(* Logix 5000 project; controller PLC_MCC1201_220AP1 vendor 1 type 14 code 164 rev 35.11; software revision 35.00; part 2 of 25 *)
(* tags used below, declared in another part *)
   N124 : DINT[414];
   N125 : DINT[414];
   N15 : DINT[1000];
   N179 : DINT[600];
   N251 : DINT[999];
   N42 : DINT[89];
   N43 : DINT[240];
   N45 : DINT[58];
   N46 : DINT[7];
   N54 : DINT[501];
   N60 : DINT[420];
   N61 : DINT[100];
   N7 : DINT[250];
   N98 : DINT[20];
   O : INT[128];
   S : INT[128];
   Status : INT;   // INT tag to retrieve Status value through GSV created during conversion
   T4 : TIMER[100];
   T51 : TIMER[13];
   TONY : ALIAS FOR B3[10].15;
   W_N7 : DINT[933];

ADD_ON_INSTRUCTION AOI_AccessArea_Logic   (* revision 1.0, vendor Bottero *)
// Help:
// (AOI_AccessArea_Logic,IN_xResetAlarm,IN_xEnableControlError,IN_xCycleON,IN_xConditionOkAccessArea,IN_xPhaseInProgressArea,IN_xExternalConditionOkToWork,IN_xSBRequestAccessAreaSelector,IN_xSBRequestAccessAreaButton,IN_xSBResetAccessArea,IN_xSBInternalResetArea,IN_xStatusDoorPH,IN_xSafetyOk,IN_xLampClock,tHMR,tAlm);
VAR_IN_OUT
   tAlm : AOI_AccessArea_Alm; {required}
   tHMR : AOI_AccessArea_HMR; {required}
END_VAR
VAR_INPUT
   IN_xConditionOkAccessArea : BOOL; {access None}
   IN_xCycleON : BOOL; {access None}
   IN_xEnableControlError : BOOL; {access None}
   IN_xLampClock : BOOL; {access None}
   IN_xPhaseInProgressArea : BOOL; {access None}
   IN_xResetAlarm : BOOL; {access None}
   IN_xSafetyOk : BOOL; {access None}
   IN_xSBInternalResetArea : BOOL; {access None}
   IN_xSBRequestAccessAreaButton : BOOL; {access None}
   IN_xSBRequestAccessAreaSelector : BOOL; {access None}
   IN_xSBResetAccessArea : BOOL; {access None}
   IN_xStatusDoorPH : BOOL; {access None}
END_VAR
VAR_OUTPUT
   OUT_xAccessAreaAccepted : BOOL; {access None}
   OUT_xAccessAreaRequest : BOOL; {access None}
   OUT_xConditionOkToWork : BOOL; {access None}
   OUT_xReqResetPhase : BOOL; {access None}
   OUT_xReqResetSafetyArea : BOOL; {access None}
   OUT_xSafetyAreaIntervened : BOOL;
   OUT_xSBLampAccessArea : BOOL;
   OUT_xSBLampInternalReset : BOOL;
   OUT_xSQOpeningDoor : BOOL;
   OUT_xStopFault : BOOL; {access None}
END_VAR
VAR_INPUT
   IN_xSAEnableResetAreaSafety : BOOL; {access None}
END_VAR
VAR
   tAOI_AccessArea_GP : AOI_AccessArea; {access None}
   ST_xConditionOkForceAccess : BOOL; {access None}
   ST_xConditionOkForRequestAccessArea : BOOL; {access None}
   ST_xErrorMutingDuringAccessArea : BOOL; {access None}
   ST_xFault : BOOL; {access None}
   ST_xInternalResetAreaRequired : BOOL; {access None}
   ST_xRequestResetPhase : BOOL; {access None}
   ST_xRequestResetSafetyArea : BOOL; {access None}
   ST_xStopFault : BOOL; {access None}
   ST_xWarning : BOOL; {access None}
   tm_ErrorMutingDuringAccessArea : TIMER; {access None}
   TMP_dAlarm : DINT; {access None}
   InitAlm : UDT_Spare32bit_Alm; {access None}
END_VAR

ROUTINE Logic   (* ladder *)
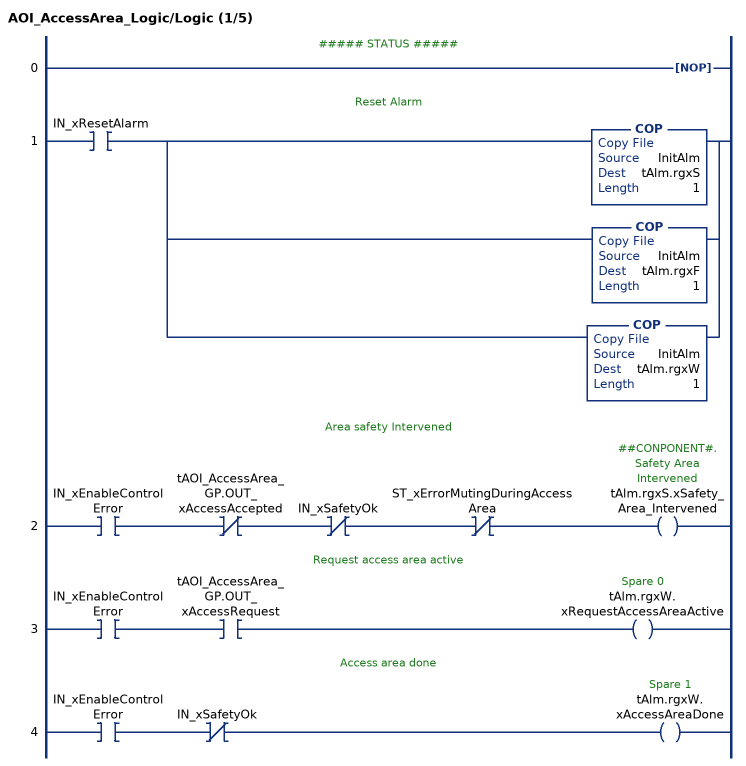
   // ##### STATUS #####
   0: NOP();
   // Reset Alarm
   1: XIC(IN_xResetAlarm)[COP(InitAlm,tAlm.rgxS,1) ,COP(InitAlm,tAlm.rgxF,1) ,COP(InitAlm,tAlm.rgxW,1) ];
   // Area safety Intervened
   2: XIC(IN_xEnableControlError)XIO(tAOI_AccessArea_GP.OUT_xAccessAccepted)XIO(IN_xSafetyOk)XIO(ST_xErrorMutingDuringAccessArea)OTE(tAlm.rgxS.xSafety_Area_Intervened);
   // Request access area active
   3: XIC(IN_xEnableControlError)XIC(tAOI_AccessArea_GP.OUT_xAccessRequest)OTE(tAlm.rgxW.xRequestAccessAreaActive);
   // Access area done
   4: XIC(IN_xEnableControlError)XIO(IN_xSafetyOk)OTE(tAlm.rgxW.xAccessAreaDone);
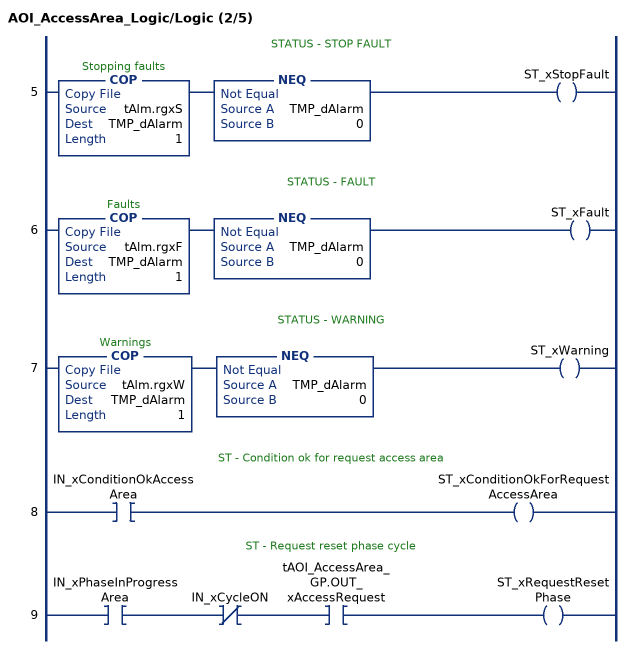
   // STATUS - STOP FAULT
   5: COP(tAlm.rgxS,TMP_dAlarm,1)NEQ(TMP_dAlarm,0)OTE(ST_xStopFault);
   // STATUS - FAULT
   6: COP(tAlm.rgxF,TMP_dAlarm,1)NEQ(TMP_dAlarm,0)OTE(ST_xFault);
   // STATUS - WARNING
   7: COP(tAlm.rgxW,TMP_dAlarm,1)NEQ(TMP_dAlarm,0)OTE(ST_xWarning);
   // ST - Condition ok for request access area
   8: XIC(IN_xConditionOkAccessArea)OTE(ST_xConditionOkForRequestAccessArea);
   // ST - Request reset phase cycle
   9: XIC(IN_xPhaseInProgressArea)XIO(IN_xCycleON)XIC(tAOI_AccessArea_GP.OUT_xAccessRequest)OTE(ST_xRequestResetPhase);
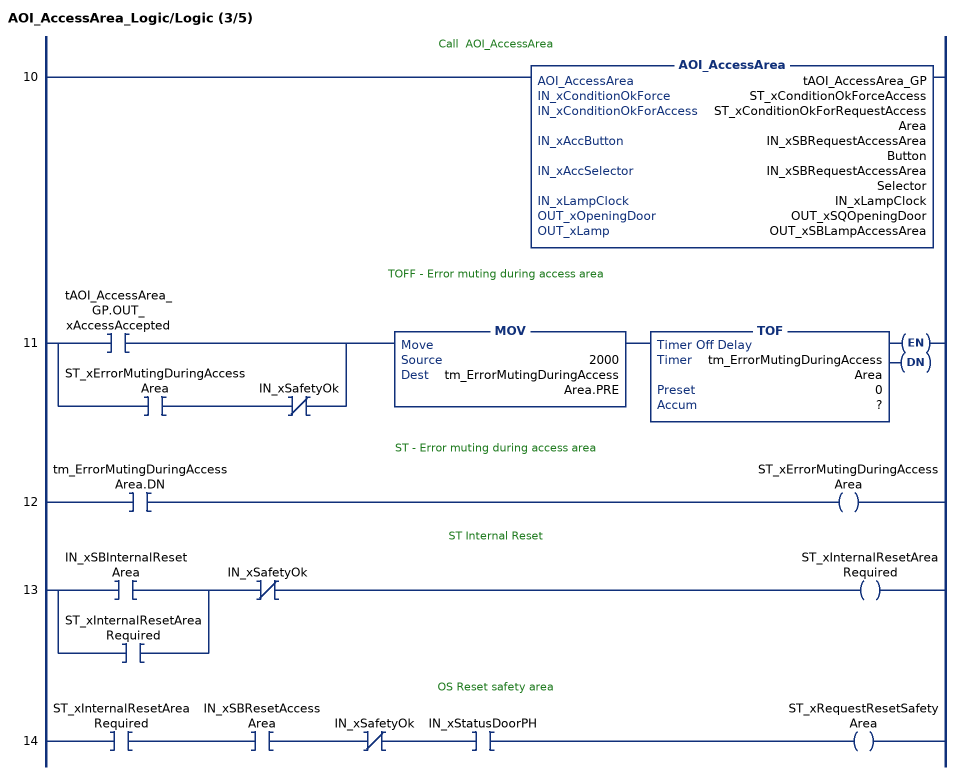
   // Call  AOI_AccessArea
   10: AOI_AccessArea(tAOI_AccessArea_GP,ST_xConditionOkForceAccess,ST_xConditionOkForRequestAccessArea,IN_xSBRequestAccessAreaButton,IN_xSBRequestAccessAreaSelector,IN_xLampClock,OUT_xSQOpeningDoor,OUT_xSBLampAccessArea);
   // TOFF - Error muting during access area
   11: [XIC(tAOI_AccessArea_GP.OUT_xAccessAccepted) ,XIC(ST_xErrorMutingDuringAccessArea) XIO(IN_xSafetyOk) ]MOV(2000,tm_ErrorMutingDuringAccessArea.PRE)TOF(tm_ErrorMutingDuringAccessArea,?,?);
   // ST - Error muting during access area
   12: XIC(tm_ErrorMutingDuringAccessArea.DN)OTE(ST_xErrorMutingDuringAccessArea);
   // ST Internal Reset
   13: [XIC(IN_xSBInternalResetArea) ,XIC(ST_xInternalResetAreaRequired) ]XIO(IN_xSafetyOk)OTE(ST_xInternalResetAreaRequired);
   // OS Reset safety area
   14: XIC(ST_xInternalResetAreaRequired)XIC(IN_xSBResetAccessArea)XIO(IN_xSafetyOk)XIC(IN_xStatusDoorPH)OTE(ST_xRequestResetSafetyArea);
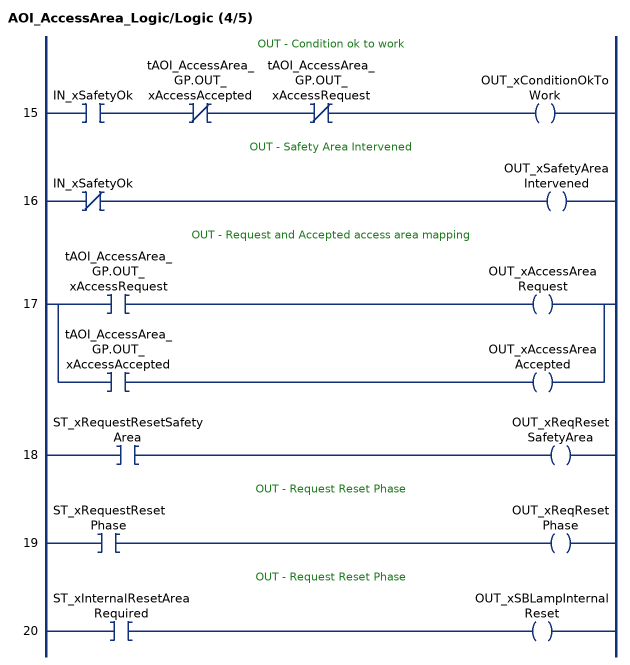
   // OUT - Condition ok to work
   15: XIC(IN_xSafetyOk)XIO(tAOI_AccessArea_GP.OUT_xAccessAccepted)XIO(tAOI_AccessArea_GP.OUT_xAccessRequest)OTE(OUT_xConditionOkToWork);
   // OUT - Safety Area Intervened
   16: XIO(IN_xSafetyOk)OTE(OUT_xSafetyAreaIntervened);
   // OUT - Request and Accepted access area mapping
   17: [XIC(tAOI_AccessArea_GP.OUT_xAccessRequest) OTE(OUT_xAccessAreaRequest) ,XIC(tAOI_AccessArea_GP.OUT_xAccessAccepted) OTE(OUT_xAccessAreaAccepted) ];
   18: XIC(ST_xRequestResetSafetyArea)OTE(OUT_xReqResetSafetyArea);
   // OUT - Request Reset Phase
   19: XIC(ST_xRequestResetPhase)OTE(OUT_xReqResetPhase);
   // OUT - Request Reset Phase
   20: XIC(ST_xInternalResetAreaRequired)OTE(OUT_xSBLampInternalReset);
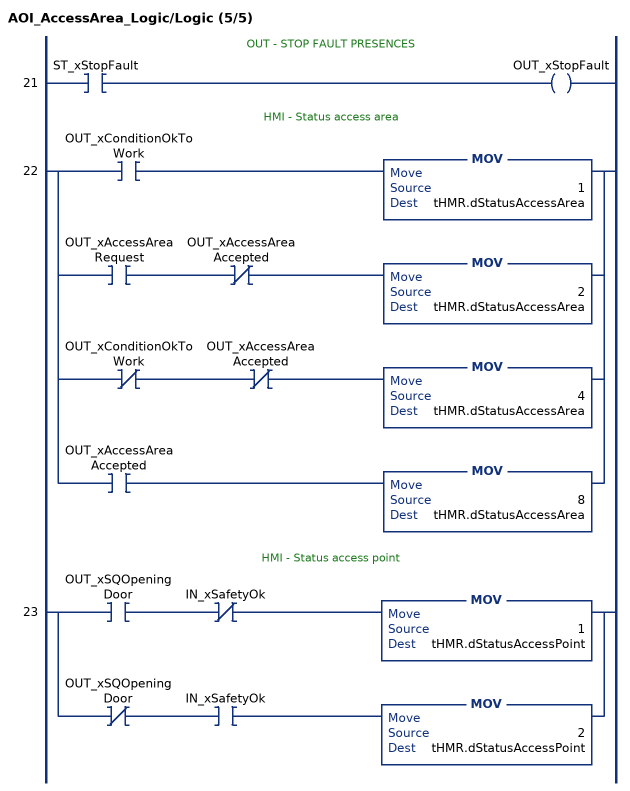
   // OUT - STOP FAULT PRESENCES
   21: XIC(ST_xStopFault)OTE(OUT_xStopFault);
   // HMI - Status access area
   22: [XIC(OUT_xConditionOkToWork) MOV(1,tHMR.dStatusAccessArea) ,XIC(OUT_xAccessAreaRequest) XIO(OUT_xAccessAreaAccepted) MOV(2,tHMR.dStatusAccessArea) ,XIO(OUT_xConditionOkToWork) XIO(OUT_xAccessAreaAccepted) MOV(4,tHMR.dStatusAccessArea) ,XIC(OUT_xAccessAreaAccepted) MOV(8,tHMR.dStatusAccessArea) ];
   // HMI - Status access point
   23: [XIC(OUT_xSQOpeningDoor) XIO(IN_xSafetyOk) MOV(1,tHMR.dStatusAccessPoint) ,XIO(OUT_xSQOpeningDoor) XIC(IN_xSafetyOk) MOV(2,tHMR.dStatusAccessPoint) ];
END_ROUTINE
END_ADD_ON_INSTRUCTION

ADD_ON_INSTRUCTION GP_AccessArea   (* revision 1.0 *)
VAR_IN_OUT
   STC : GP_AccessArea_STC; {required}
END_VAR
VAR_INPUT
   IN_xAccSelector : BOOL; {access None, required}
   IN_xAccButton : BOOL; {access None, required}
   IN_xConditionOkAccess : BOOL; {access None, required}
   IN_xConditionOkForcedAccess : BOOL; {access None, required}
   IN_xLampClock : BOOL; {access None, required}
END_VAR
VAR_OUTPUT
   OUT_xOpeningDoor : BOOL; {access None}
   OUT_xLamp : BOOL; {access None, required}
END_VAR

ROUTINE Logic   (* ladder *)
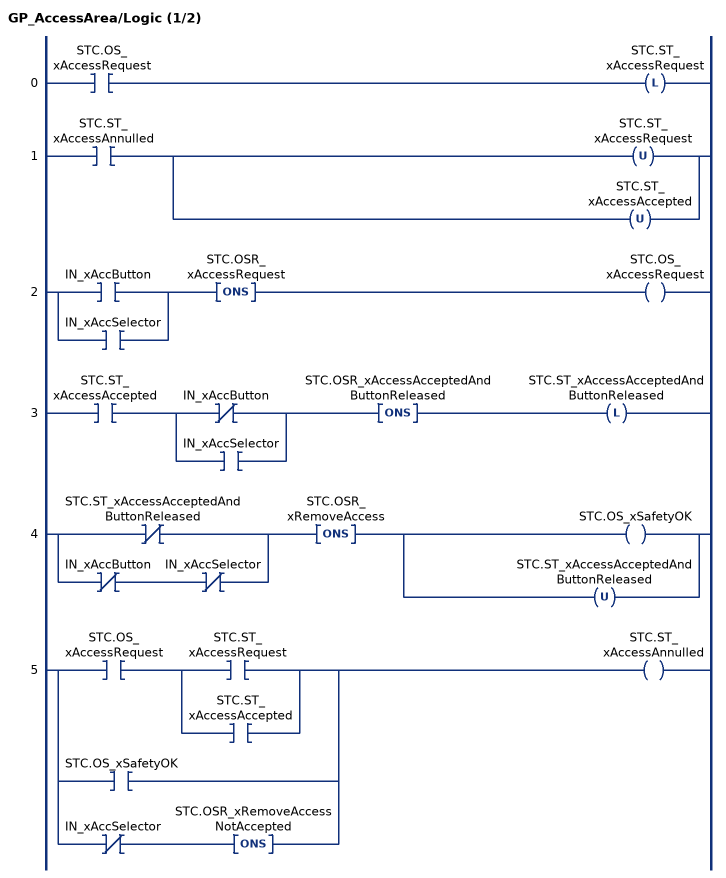
   0: XIC(STC.OS_xAccessRequest)OTL(STC.ST_xAccessRequest);
   1: XIC(STC.ST_xAccessAnnulled)[OTU(STC.ST_xAccessRequest) ,OTU(STC.ST_xAccessAccepted) ];
   2: [XIC(IN_xAccButton) ,XIC(IN_xAccSelector) ]ONS(STC.OSR_xAccessRequest)OTE(STC.OS_xAccessRequest);
   3: XIC(STC.ST_xAccessAccepted)[XIO(IN_xAccButton) ,XIC(IN_xAccSelector) ]ONS(STC.OSR_xAccessAcceptedAndButtonReleased)OTL(STC.ST_xAccessAcceptedAndButtonReleased);
   4: [XIO(STC.ST_xAccessAcceptedAndButtonReleased) ,XIO(IN_xAccButton) XIO(IN_xAccSelector) ]ONS(STC.OSR_xRemoveAccess)[OTE(STC.OS_xSafetyOK) ,OTU(STC.ST_xAccessAcceptedAndButtonReleased) ];
   5: [XIC(STC.OS_xAccessRequest) [XIC(STC.ST_xAccessRequest) ,XIC(STC.ST_xAccessAccepted) ] ,XIC(STC.OS_xSafetyOK) ,XIO(IN_xAccSelector) ONS(STC.OSR_xRemoveAccessNotAccepted) ]OTE(STC.ST_xAccessAnnulled);
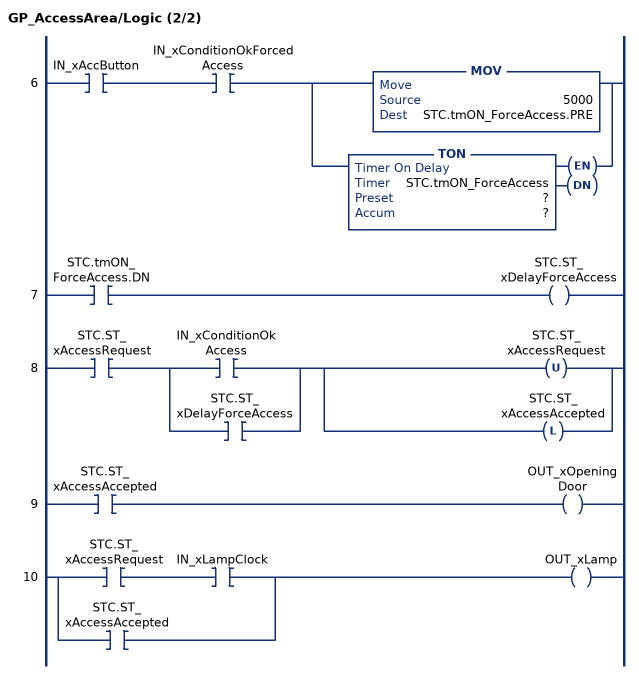
   6: XIC(IN_xAccButton)XIC(IN_xConditionOkForcedAccess)[MOV(5000,STC.tmON_ForceAccess.PRE) ,TON(STC.tmON_ForceAccess,?,?) ];
   7: XIC(STC.tmON_ForceAccess.DN)OTE(STC.ST_xDelayForceAccess);
   8: XIC(STC.ST_xAccessRequest)[XIC(IN_xConditionOkAccess) ,XIC(STC.ST_xDelayForceAccess) ][OTU(STC.ST_xAccessRequest) ,OTL(STC.ST_xAccessAccepted) ];
   9: XIC(STC.ST_xAccessAccepted)OTE(OUT_xOpeningDoor);
   10: [XIC(STC.ST_xAccessRequest) XIC(IN_xLampClock) ,XIC(STC.ST_xAccessAccepted) ]OTE(OUT_xLamp);
END_ROUTINE
END_ADD_ON_INSTRUCTION

ADD_ON_INSTRUCTION GP_NetworkDiag   (* revision 1.0 *)
VAR_IN_OUT
   IN_OB_Initialize : GP_OB_Initialize; {required}
   IN_ModuleName : MODULE; {required}   // Module name
   OUT_tModuleInfo : GP_NetworkDiag_v1; {required}   // Module info
END_VAR
VAR
   TMP_xFaulted : BOOL; {access None}
   TMP_xConnected : BOOL; {access None}
END_VAR

ROUTINE Logic   (* structured text *)
   //Initialize
   TMP_xConnected:=0;
   TMP_xFaulted:=0;
   
   //Get system info from module
   gsv(Module,IN_ModuleName,EntryStatus,OUT_tModuleInfo.dEntryStatus);
   gsv(Module,IN_ModuleName,FaultCode,OUT_tModuleInfo.dFaultCode);
   gsv(Module,IN_ModuleName,FaultInfo,OUT_tModuleInfo.dFaultInfo);
   gsv(Module,IN_ModuleName,Instance,OUT_tModuleInfo.dInstance);
   
   CASE OUT_tModuleInfo.dEntryStatus OF
   	16#0000:(*Standby: the controller is powering up.*)
    			TMP_xFaulted:= IN_OB_Initialize.OUT_xClock_800ms;
   
   	16#1000:(*Faulted: any of the MODULE object’s connections to the associated module fail.
   			This value should not be used to determine if the module failed because the MODULE
   			object leaves this state periodically when trying to reconnect to the module.
   			Instead, test for Running state (16#4000). Check for FaultCode not equal to 0 to determine if a module is faulted.
   			When Faulted, the FaultCode and FaultInfo attributes are valid until the fault condition is corrected.*)
    			TMP_xConnected:= IN_OB_Initialize.OUT_xClock_1s;
   			TMP_xFaulted:= 1;
   
   	16#2000:(*Validating: the MODULE object is verifying MODULE object integrity prior to establishing connections to the module.*)
    			TMP_xConnected:= IN_OB_Initialize.OUT_xClock_400ms;
   
   	16#3000:(*Connecting: the MODULE object is initiating connections to the module.*)
   			TMP_xConnected:= IN_OB_Initialize.OUT_xClock_400ms;
   
   	16#4000:(*Running: all connections to the module are established and data is successfully transferring.*)
    			TMP_xConnected:= 1;
   
   	16#5000:(*Shutting down: the MODULE object is in the process of shutting down all connections to the module.*)
   			TMP_xConnected:= IN_OB_Initialize.OUT_xClock_1s;
   
   	16#6000:(*Inhibited: the MODULE object is inhibited (the inhibit bit in the Mode attribute is set).*)
    			TMP_xConnected:= IN_OB_Initialize.OUT_xClock_1s;
   
   	16#7000:(*Waiting: the parent MODULE object upon which this MODULE object depends is not running*)
   			TMP_xConnected:= IN_OB_Initialize.OUT_xClock_1s;
   
   	16#9000:(*FirmwareUpdating: Firmware supervisor is attempting to flash the module. *)
    			TMP_xConnected:= IN_OB_Initialize.OUT_xClock_800ms;
   
   	16#A000:(*Configuring: Controller is downloading configuration to the module.
   			Either ?forward open? or (ADC) download occur during this state.*)
   			TMP_xConnected:= IN_OB_Initialize.OUT_xClock_800ms;
   END_CASE;
   
   IF OUT_tModuleInfo.dFaultCode<>0 THEN
   	TMP_xFaulted:= 1;
   	TMP_xConnected:= 0;
   END_IF;
   
   //Save status bit
   OUT_tModuleInfo.xConnected:=TMP_xConnected;
   OUT_tModuleInfo.xFaulted:=TMP_xFaulted;
   
   
   
   
   
   
   
   
   
   
   
   
   
   
   
   
   
   
   
   
END_ROUTINE
END_ADD_ON_INSTRUCTION

ADD_ON_INSTRUCTION GP_OB_Initialize   (* revision 1.0 *)
VAR_IN_OUT
   STC : GP_OB_Initialize_STC; {required}
END_VAR
VAR_INPUT
   IN_xInitialize : BOOL; {access None, required}   // Initialize values (Restart call)
END_VAR
VAR_OUTPUT
   OUT_dExecutionTime_ms : DINT; {access None}   // OB Execution time [ms]
   OUT_dMinExecutionTime_ms : DINT; {access None}   // OB Minimum execution time [ms]
   OUT_dMaxExecutionTime_ms : DINT; {access None}   // OB Maximum execution time [ms]
   OUT_xOs_100ms : BOOL; {access None}   // OS each 100ms
   OUT_xOs_200ms : BOOL; {access None}   // OS each 200ms
   OUT_xOs_400ms : BOOL; {access None}   // OS each 400ms
   OUT_xOs_500ms : BOOL; {access None}   // OS each 500ms
   OUT_xOs_800ms : BOOL; {access None}   // OS each 800ms
   OUT_xOs_1s : BOOL; {access None}   // OS each 1s
   OUT_xOs_2s : BOOL; {access None}   // OS each 2s
   OUT_xOs_5s : BOOL; {access None}   // OS each 5s
   OUT_xOs_10s : BOOL; {access None}   // OS each 10s
   OUT_xOs_30s : BOOL; {access None}   // OS each 30s
   OUT_xOs_1min : BOOL; {access None}   // OS each 1min
   OUT_xOs_2min : BOOL; {access None}   // OS each 2min
   OUT_xOs_10min : BOOL; {access None}   // OS each 10min
   OUT_xOs_30min : BOOL; {access None}   // OS each 30min
   OUT_xOs_1h : BOOL; {access None}   // OS each 1h
   OUT_xClock_100ms : BOOL; {access None}   // Clock 100ms
   OUT_xClock_200ms : BOOL; {access None}   // Clock 200ms
   OUT_xClock_400ms : BOOL; {access None}   // Clock 400ms
   OUT_xClock_500ms : BOOL; {access None}   // Clock 500ms
   OUT_xClock_800ms : BOOL; {access None}   // Clock 800ms
   OUT_xClock_1s : BOOL; {access None}   // Clock 1s
   OUT_xClock_2s : BOOL; {access None}   // Clock 2s
   OUT_xClock_5s : BOOL; {access None}   // Clock 5s
   OUT_xClock_10s : BOOL; {access None}   // Clock 10s
   OUT_xClock_30s : BOOL; {access None}   // Clock 30s
   OUT_xClock_1min : BOOL; {access None}   // Clock 1min
   OUT_xClock_2min : BOOL; {access None}   // Clock 2min
   OUT_xClock_10min : BOOL; {access None}   // Clock 10min
   OUT_xClock_30min : BOOL; {access None}   // Clock 30min
   OUT_xClock_1h : BOOL; {access None}   // Clock 1h
   OUT_xDebugOFF : BOOL; {access None}
   OUT_xDebugON : BOOL; {access None}
END_VAR
VAR
   CONST_DMAX_INT : DINT; {access None}
   CONST_DTICK_1H : DINT; {access None}
   CONST_DTICK_30MIN : DINT; {access None}
   CONST_DTICK_10MIN : DINT; {access None}
   CONST_DTICK_2MIN : DINT; {access None}
   CONST_DTICK_1MIN : DINT; {access None}
   CONST_DTICK_30S : DINT; {access None}
   CONST_DTICK_10S : DINT; {access None}
   CONST_DTICK_5S : DINT; {access None}
   CONST_DTICK_2S : DINT; {access None}
   CONST_DTICK_1S : DINT; {access None}
   CONST_DTICK_800MS : DINT; {access None}
   CONST_DTICK_500MS : DINT; {access None}
   CONST_DTICK_400MS : DINT; {access None}
   CONST_DTICK_200MS : DINT; {access None}
   CONST_DTICK_100MS : DINT; {access None}
   TMP_rlActualExecutionTimeRound : REAL; {access None}   // Rounded execution time [ms]
   TMP_rlActualExecutionTime : REAL; {access None}   // ActualExecutionTime [ms]
END_VAR

ROUTINE Logic   (* structured text *)
   //Costants
   CONST_DTICK_100MS:=100;
   CONST_DTICK_200MS:=200;
   CONST_DTICK_400MS:=400;
   CONST_DTICK_500MS:=500;
   CONST_DTICK_800MS:=800;
   CONST_DTICK_1S:=1000;
   CONST_DTICK_2S:=2000;
   CONST_DTICK_5S:=5000;
   CONST_DTICK_10S:=10000;
   CONST_DTICK_30S:=30000;
   CONST_DTICK_1MIN:=60000;
   CONST_DTICK_2MIN:=120000;
   CONST_DTICK_10MIN:=600000;
   CONST_DTICK_30MIN:=1800000;
   CONST_DTICK_1H:=86400000;
   CONST_DMAX_INT:=16#7FFFFFFF;
   OUT_xDebugOFF:=0;
   OUT_xDebugON:=1;
   
   //Initialize OS bits
   OUT_xOs_100ms := 0;
   OUT_xOs_200ms := 0;
   OUT_xOs_400ms := 0;
   OUT_xOs_500ms := 0;
   OUT_xOs_800ms := 0;
   OUT_xOs_1s := 0;
   OUT_xOs_2s := 0;
   OUT_xOs_5s := 0;
   OUT_xOs_10s := 0;
   OUT_xOs_30s := 0;
   OUT_xOs_1min := 0;
   OUT_xOs_2min := 0;
   OUT_xOs_10min := 0;
   OUT_xOs_30min := 0;
   OUT_xOs_1h := 0;
   
   //Take the start execution time from the CPU
   gsv(Task,THIS,StartTime,STC.lwStartTime[0]);
   
   //Initialize FB execution
   IF IN_xInitialize THEN
   
   	IN_xInitialize := 0;
   	OUT_dExecutionTime_ms := 0;
   	OUT_dMinExecutionTime_ms := CONST_DMAX_INT;
   	OUT_dMaxExecutionTime_ms := 0;
   	OUT_xClock_100ms := 0;
   	OUT_xClock_200ms := 0;
   	OUT_xClock_400ms := 0;
   	OUT_xClock_500ms := 0;
   	OUT_xClock_800ms := 0;
   	OUT_xClock_1s := 0;
   	OUT_xClock_2s := 0;
   	OUT_xClock_5s := 0;
   	OUT_xClock_10s := 0;
   	OUT_xClock_30s := 0;
   	OUT_xClock_1min := 0;
   	OUT_xClock_2min := 0;
   	OUT_xClock_10min := 0;
   	OUT_xClock_30min := 0;
   	OUT_xClock_1h := 0;
   
   	STC.dElapsed_100ms_ms := 0;
   	STC.dElapsed_200ms_ms := 0;
   	STC.dElapsed_400ms_ms := 0;
   	STC.dElapsed_500ms_ms := 0;
   	STC.dElapsed_800ms_ms := 0;
   	STC.dElapsed_1s_ms := 0;
   	STC.dElapsed_2s_ms := 0;
   	STC.dElapsed_5s_ms := 0;
   	STC.dElapsed_10s_ms := 0;
   	STC.dElapsed_30s_ms := 0;
   	STC.dElapsed_1min_ms := 0;
   	STC.dElapsed_2min_ms := 0;
   	STC.dElapsed_10min_ms := 0;
   	STC.dElapsed_30min_ms := 0;
   	STC.dElapsed_1h_ms := 0;
   
   	STC.lwOldStartTime[0] := STC.lwStartTime[0];
   	STC.lwOldStartTime[1] := STC.lwStartTime[1];
   
   END_IF;
   
   //***** CALCULATE OB EXECUTION TIME *****
   STC.dlLastExecValue_us := STC.lwStartTime[0] - STC.lwOldStartTime[0];
   STC.lwOldStartTime[0] := STC.lwStartTime[0];
   STC.lwOldStartTime[1] := STC.lwStartTime[1];
   //Convert from [us] to [ms]
   TMP_rlActualExecutionTime := STC.dlLastExecValue_us / 1000.0;
   //Add the reminder of the last cycle
   TMP_rlActualExecutionTime := TMP_rlActualExecutionTime + STC.rReminder_ms;
   //Calculate the rounded value
   TMP_rlActualExecutionTimeRound:= trunc(TMP_rlActualExecutionTime + 0.5);
   OUT_dExecutionTime_ms := trunc(TMP_rlActualExecutionTime + 0.5);
   //Save the reminder for the next cycle
   STC.rReminder_ms := TMP_rlActualExecutionTime - TMP_rlActualExecutionTimeRound;
   
   //Save the maximum scan value
   IF OUT_dExecutionTime_ms > OUT_dMaxExecutionTime_ms THEN
   	OUT_dMaxExecutionTime_ms := OUT_dExecutionTime_ms;
   END_IF;
   
   //Save the minimum scan value
   IF OUT_dExecutionTime_ms < OUT_dMinExecutionTime_ms THEN
   	OUT_dMinExecutionTime_ms := OUT_dExecutionTime_ms;
   END_IF;
   
   //***** CALCULATE SERVICES CLOCK *****
   
   //Increment counters for each clock
   STC.dElapsed_100ms_ms := STC.dElapsed_100ms_ms + OUT_dExecutionTime_ms;
   STC.dElapsed_200ms_ms := STC.dElapsed_200ms_ms + OUT_dExecutionTime_ms;
   STC.dElapsed_400ms_ms := STC.dElapsed_400ms_ms + OUT_dExecutionTime_ms;
   STC.dElapsed_500ms_ms := STC.dElapsed_500ms_ms + OUT_dExecutionTime_ms;
   STC.dElapsed_800ms_ms := STC.dElapsed_800ms_ms + OUT_dExecutionTime_ms;
   STC.dElapsed_1s_ms := STC.dElapsed_1s_ms + OUT_dExecutionTime_ms;
   STC.dElapsed_2s_ms := STC.dElapsed_2s_ms + OUT_dExecutionTime_ms;
   STC.dElapsed_5s_ms := STC.dElapsed_5s_ms + OUT_dExecutionTime_ms;
   STC.dElapsed_10s_ms := STC.dElapsed_10s_ms + OUT_dExecutionTime_ms;
   STC.dElapsed_30s_ms := STC.dElapsed_30s_ms + OUT_dExecutionTime_ms;
   STC.dElapsed_1min_ms := STC.dElapsed_1min_ms + OUT_dExecutionTime_ms;
   STC.dElapsed_2min_ms := STC.dElapsed_2min_ms + OUT_dExecutionTime_ms;
   STC.dElapsed_10min_ms := STC.dElapsed_10min_ms + OUT_dExecutionTime_ms;
   STC.dElapsed_30min_ms := STC.dElapsed_30min_ms + OUT_dExecutionTime_ms;
   STC.dElapsed_1h_ms := STC.dElapsed_1h_ms + OUT_dExecutionTime_ms;
   
   //Calculate the 100ms
   IF STC.dElapsed_100ms_ms >= CONST_DTICK_100MS THEN
   	STC.dElapsed_100ms_ms := STC.dElapsed_100ms_ms - CONST_DTICK_100MS;
   
   	OUT_xOs_100ms := 1;
   
   	IF NOT(OUT_xClock_100ms) THEN
   		OUT_xClock_100ms := 1;
   	ELSE
   		OUT_xClock_100ms := 0;
   	END_IF;
   END_IF;
   
   //Calculate the 200ms
   IF STC.dElapsed_200ms_ms >= CONST_DTICK_200MS THEN
   	STC.dElapsed_200ms_ms := STC.dElapsed_200ms_ms - CONST_DTICK_200MS;
   
   	OUT_xOs_200ms := 1;
   
   	IF NOT(OUT_xClock_200ms) THEN
   		OUT_xClock_200ms := 1;
   	ELSE
   		OUT_xClock_200ms := 0;
   	END_IF;
   END_IF;
   
   //Calculate the 400ms
   IF STC.dElapsed_400ms_ms >= CONST_DTICK_400MS THEN
   	STC.dElapsed_400ms_ms := STC.dElapsed_400ms_ms - CONST_DTICK_400MS;
   
   	OUT_xOs_400ms := 1;
   
   	IF NOT(OUT_xClock_400ms) THEN
   		OUT_xClock_400ms := 1;
   	ELSE
   		OUT_xClock_400ms := 0;
   	END_IF;
   END_IF;
   
   //Calculate the 500ms
   IF STC.dElapsed_500ms_ms >= CONST_DTICK_500MS THEN
   	STC.dElapsed_500ms_ms := STC.dElapsed_500ms_ms - CONST_DTICK_500MS;
   
   	OUT_xOs_500ms := 1;
   
   	IF NOT(OUT_xClock_500ms) THEN
   		OUT_xClock_500ms := 1;
   	ELSE
   		OUT_xClock_500ms := 0;
   	END_IF;
   END_IF;
   
   //Calculate the 800ms
   IF STC.dElapsed_800ms_ms >= CONST_DTICK_800MS THEN
   	STC.dElapsed_800ms_ms := STC.dElapsed_800ms_ms - CONST_DTICK_800MS;
   
   	OUT_xOs_800ms := 1;
   
   	IF NOT(OUT_xClock_800ms) THEN
   		OUT_xClock_800ms := 1;
   	ELSE
   		OUT_xClock_800ms := 0;
   	END_IF;
   END_IF;
   
   //Calculate the 1s
   IF STC.dElapsed_1s_ms >= CONST_DTICK_1S THEN
   	STC.dElapsed_1s_ms := STC.dElapsed_1s_ms - CONST_DTICK_1S;
   
   	OUT_xOs_1s := 1;
   
   	IF NOT(OUT_xClock_1s) THEN
   		OUT_xClock_1s := 1;
   	ELSE
   		OUT_xClock_1s := 0;
   	END_IF;
   END_IF;
   
   //Calculate the 2s
   IF STC.dElapsed_2s_ms >= CONST_DTICK_2S THEN
   	STC.dElapsed_2s_ms := STC.dElapsed_2s_ms - CONST_DTICK_2S;
   
   	OUT_xOs_2s := 1;
   
   	IF NOT(OUT_xClock_2s) THEN
   		OUT_xClock_2s := 1;
   	ELSE
   		OUT_xClock_2s := 0;
   	END_IF;
   END_IF;
   
   //Calculate the 5s
   IF STC.dElapsed_5s_ms >= CONST_DTICK_5S THEN
   	STC.dElapsed_5s_ms := STC.dElapsed_5s_ms - CONST_DTICK_5S;
   
   	OUT_xOs_5s := 1;
   
   	IF NOT(OUT_xClock_5s) THEN
   		OUT_xClock_5s := 1;
   	ELSE
   		OUT_xClock_5s := 0;
   	END_IF;
   END_IF;
   
   //Calculate the 10s
   IF STC.dElapsed_10s_ms >= CONST_DTICK_10S THEN
   	STC.dElapsed_10s_ms := STC.dElapsed_10s_ms - CONST_DTICK_10S;
   
   	OUT_xOs_10s := 1;
   
   	IF NOT(OUT_xClock_10s) THEN
   		OUT_xClock_10s := 1;
   	ELSE
   		OUT_xClock_10s := 0;
   	END_IF;
   END_IF;
   
   //Calculate the 30s
   IF STC.dElapsed_30s_ms >= CONST_DTICK_30S THEN
   	STC.dElapsed_30s_ms := STC.dElapsed_30s_ms - CONST_DTICK_30S;
   
   	OUT_xOs_30s := 1;
   
   	IF NOT(OUT_xClock_30s) THEN
   		OUT_xClock_30s := 1;
   	ELSE
   		OUT_xClock_30s := 0;
   	END_IF;
   END_IF;
   
   //Calculate the 1min
   IF STC.dElapsed_1min_ms >= CONST_DTICK_1MIN THEN
   	STC.dElapsed_1min_ms := STC.dElapsed_1min_ms - CONST_DTICK_1MIN;
   
   	OUT_xOs_1min := 1;
   
   	IF NOT(OUT_xClock_1min) THEN
   		OUT_xClock_1min := 1;
   	ELSE
   		OUT_xClock_1min := 0;
   	END_IF;
   END_IF;
   
   //Calculate the 2min
   IF STC.dElapsed_2min_ms >= CONST_DTICK_2MIN THEN
   	STC.dElapsed_2min_ms := STC.dElapsed_2min_ms - CONST_DTICK_2MIN;
   
   	OUT_xOs_2min := 1;
   
   	IF NOT(OUT_xClock_2min) THEN
   		OUT_xClock_2min := 1;
   	ELSE
   		OUT_xClock_2min := 0;
   	END_IF;
   END_IF;
   
   //Calculate the 10min
   IF STC.dElapsed_10min_ms >= CONST_DTICK_10MIN THEN
   	STC.dElapsed_10min_ms := STC.dElapsed_10min_ms - CONST_DTICK_10MIN;
   
   	OUT_xOs_10min := 1;
   
   	IF NOT(OUT_xClock_10min) THEN
   		OUT_xClock_10min := 1;
   	ELSE
   		OUT_xClock_10min := 0;
   	END_IF;
   END_IF;
   
   //Calculate the 30min
   IF STC.dElapsed_30min_ms >= CONST_DTICK_30MIN THEN
   	STC.dElapsed_30min_ms := STC.dElapsed_30min_ms - CONST_DTICK_30MIN;
   
   	OUT_xOs_30min := 1;
   
   	IF NOT(OUT_xClock_30min) THEN
   		OUT_xClock_30min := 1;
   	ELSE
   		OUT_xClock_30min := 0;
   	END_IF;
   END_IF;
   
   //Calculate the 1h
   IF STC.dElapsed_1h_ms >= CONST_DTICK_1H THEN
   	STC.dElapsed_1h_ms := STC.dElapsed_1h_ms - CONST_DTICK_1H;
   
   	OUT_xOs_1h := 1;
   
   	IF NOT(OUT_xClock_1h) THEN
   		OUT_xClock_1h := 1;
   	ELSE
   		OUT_xClock_1h := 0;
   	END_IF;
   END_IF;
END_ROUTINE
END_ADD_ON_INSTRUCTION

ADD_ON_INSTRUCTION GP_RibbonTracking_GetRibbonData   (* revision 1.0 *)
VAR_INPUT
   INP_dMachinePositionFromSnap_cmm : DINT; {required}   // Machine position from snaproll [mm/100]
   INP_dOffsetBreakUpstream_cmm : DINT; {required}   // Offset upstream glass break [mm/100]
   INP_dOffsetBreakDownstream_cmm : DINT; {required}   // Offset downstream glass break [mm/100]
END_VAR
VAR_IN_OUT
   INO_tRibbonData : DATA_TRACKING_RIBBON; {required}   // Ribbon tracking array
END_VAR
VAR_OUTPUT
   OUT_dGrossWidth_cmm : DINT; {visible}   // Gross width [mm/100]
   OUT_dNetWidth_cmm : DINT; {visible}   // Net width [mm/100]
   OUT_dGrossWander_cmm : DINT; {visible}   // Gross wander [mm/100]
   OUT_dNetWander_cmm : DINT; {visible}   // Net wander [mm/100]
   OUT_dBreakMask : DINT; {visible}   // Break mask [Mask]
END_VAR
VAR
   TMP_dIndex : DINT; {access None}
   TMP_tRibbon : DATA_TRACKING_RIBBON_DETAILS; {access None}
   TMP_dIndexEnd : DINT; {access None}
   TMP_dIndexStart : DINT; {access None}
   TMP_dBreak : DINT; {access None}
END_VAR

ROUTINE Logic   (* structured text *)
   
   TMP_dIndexStart := (INP_dMachinePositionFromSnap_cmm - INP_dOffsetBreakUpstream_cmm) / INO_tRibbonData.dStepAdvancement_cmm;
   TMP_dIndexEnd := (INP_dMachinePositionFromSnap_cmm + INP_dOffsetBreakDownstream_cmm) / INO_tRibbonData.dStepAdvancement_cmm;
   
   //Update the data in that position
   INO_tRibbonData.dOperationInProgress := INO_tRibbonData.dOperationInProgress + 1;
   
   TMP_dBreak := 0;
   
   FOR TMP_dIndex := TMP_dIndexStart TO TMP_dIndexEnd DO
   
   	IF INO_tRibbonData.rgtRibbons[TMP_dIndex].rgxGlassBreak <> 0 THEN
   		TMP_dBreak := INO_tRibbonData.rgtRibbons[TMP_dIndex].rgxGlassBreak;
   	END_IF;
   
   END_FOR;
   
   //Find the correct position
   TMP_dIndex := INP_dMachinePositionFromSnap_cmm / INO_tRibbonData.dStepAdvancement_cmm;
   
   COP(INO_tRibbonData.rgtRibbons[TMP_dIndex], TMP_tRibbon, 1);
   
   INO_tRibbonData.dOperationInProgress := INO_tRibbonData.dOperationInProgress - 1;
   
   //Move the data on the out information
   OUT_dGrossWander_cmm := TMP_tRibbon.dGrossWander_cmm;
   OUT_dGrossWidth_cmm := TMP_tRibbon.dGrossRibbonWidth_cmm;
   OUT_dNetWander_cmm :=  TMP_tRibbon.dNetWander_cmm;
   OUT_dNetWidth_cmm := TMP_tRibbon.dNetRibbonWidth_cmm ;
   OUT_dBreakMask := TMP_dBreak;
   
END_ROUTINE
END_ADD_ON_INSTRUCTION

ADD_ON_INSTRUCTION GP_RibbonTracking_UpdateGlassBreak   (* revision 1.0 *)
VAR_INPUT
   INP_dMachinePositionFromSnap_cmm : DINT; {required}   // Machine position from snaproll [mm/100]
   INP_dBreakMask : DINT; {required}   // Break mask [Mask]
END_VAR
VAR_IN_OUT
   INO_tRibbonData : DATA_TRACKING_RIBBON; {required}   // Ribbon tracking array
END_VAR
VAR
   TMP_dIndex : DINT; {access None}
END_VAR

ROUTINE Logic   (* structured text *)
   //Find the correct position
   TMP_dIndex := INP_dMachinePositionFromSnap_cmm / INO_tRibbonData.dStepAdvancement_cmm;
   
   //Update the data in that position
   INO_tRibbonData.rgtRibbons[TMP_dIndex].rgxGlassBreak := INP_dBreakMask;
   
END_ROUTINE
END_ADD_ON_INSTRUCTION
